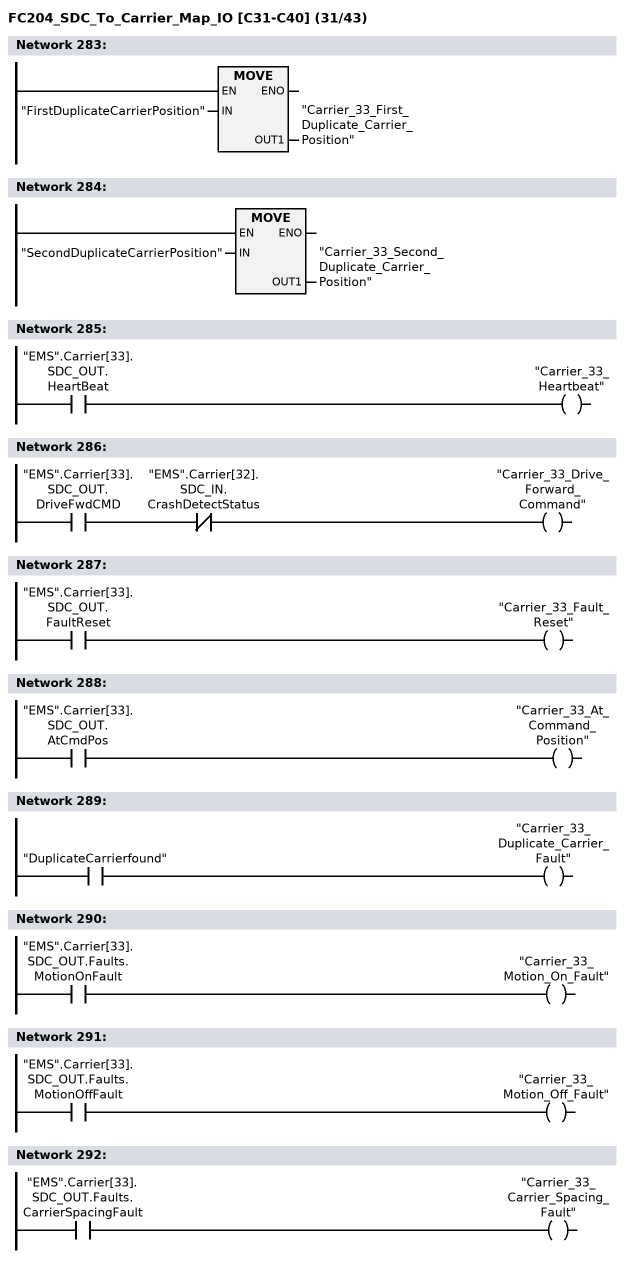
   RUNG wire#powerrail
      Move(in := "FirstDuplicateCarrierPosition", out1 => "Carrier_33_First_Duplicate_Carrier_Position")
   END_RUNG
   // the same network as SCL:
   "Carrier_33_First_Duplicate_Carrier_Position" := "FirstDuplicateCarrierPosition";
END_REGION

REGION Network 284
   RUNG wire#powerrail
      Move(in := "SecondDuplicateCarrierPosition", out1 => "Carrier_33_Second_Duplicate_Carrier_Position")
   END_RUNG
   // the same network as SCL:
   "Carrier_33_Second_Duplicate_Carrier_Position" := "SecondDuplicateCarrierPosition";
END_REGION

REGION Network 285
   RUNG wire#powerrail
      Contact( "EMS".Carrier[33].SDC_OUT.HeartBeat )
      Coil( "Carrier_33_Heartbeat" )
   END_RUNG
   // the same network as SCL:
   "Carrier_33_Heartbeat" := "EMS".Carrier[33].SDC_OUT.HeartBeat;
END_REGION

REGION Network 286
   RUNG wire#powerrail
      Contact( "EMS".Carrier[33].SDC_OUT.DriveFwdCMD )
      I_Contact( "EMS".Carrier[32].SDC_IN.CrashDetectStatus )
      Coil( "Carrier_33_Drive_Forward_Command" )
   END_RUNG
   // the same network as SCL:
   "Carrier_33_Drive_Forward_Command" := "EMS".Carrier[33].SDC_OUT.DriveFwdCMD AND NOT "EMS".Carrier[32].SDC_IN.CrashDetectStatus;
END_REGION

REGION Network 287
   RUNG wire#powerrail
      Contact( "EMS".Carrier[33].SDC_OUT.FaultReset )
      Coil( "Carrier_33_Fault_Reset" )
   END_RUNG
   // the same network as SCL:
   "Carrier_33_Fault_Reset" := "EMS".Carrier[33].SDC_OUT.FaultReset;
END_REGION

REGION Network 288
   RUNG wire#powerrail
      Contact( "EMS".Carrier[33].SDC_OUT.AtCmdPos )
      Coil( "Carrier_33_At_Command_Position" )
   END_RUNG
   // the same network as SCL:
   "Carrier_33_At_Command_Position" := "EMS".Carrier[33].SDC_OUT.AtCmdPos;
END_REGION

REGION Network 289
   RUNG wire#powerrail
      Contact( "DuplicateCarrierfound" )
      Coil( "Carrier_33_Duplicate_Carrier_Fault" )
   END_RUNG
   // the same network as SCL:
   "Carrier_33_Duplicate_Carrier_Fault" := "DuplicateCarrierfound";
END_REGION

REGION Network 290
   RUNG wire#powerrail
      Contact( "EMS".Carrier[33].SDC_OUT.Faults.MotionOnFault )
      Coil( "Carrier_33_Motion_On_Fault" )
   END_RUNG
   // the same network as SCL:
   "Carrier_33_Motion_On_Fault" := "EMS".Carrier[33].SDC_OUT.Faults.MotionOnFault;
END_REGION

REGION Network 291
   RUNG wire#powerrail
      Contact( "EMS".Carrier[33].SDC_OUT.Faults.MotionOffFault )
      Coil( "Carrier_33_Motion_Off_Fault" )
   END_RUNG
   // the same network as SCL:
   "Carrier_33_Motion_Off_Fault" := "EMS".Carrier[33].SDC_OUT.Faults.MotionOffFault;
END_REGION

REGION Network 292
   RUNG wire#powerrail
      Contact( "EMS".Carrier[33].SDC_OUT.Faults.CarrierSpacingFault )
      Coil( "Carrier_33_Carrier_Spacing_Fault" )
   END_RUNG
   // the same network as SCL:
   "Carrier_33_Carrier_Spacing_Fault" := "EMS".Carrier[33].SDC_OUT.Faults.CarrierSpacingFault;
END_REGION

REGION Network 293
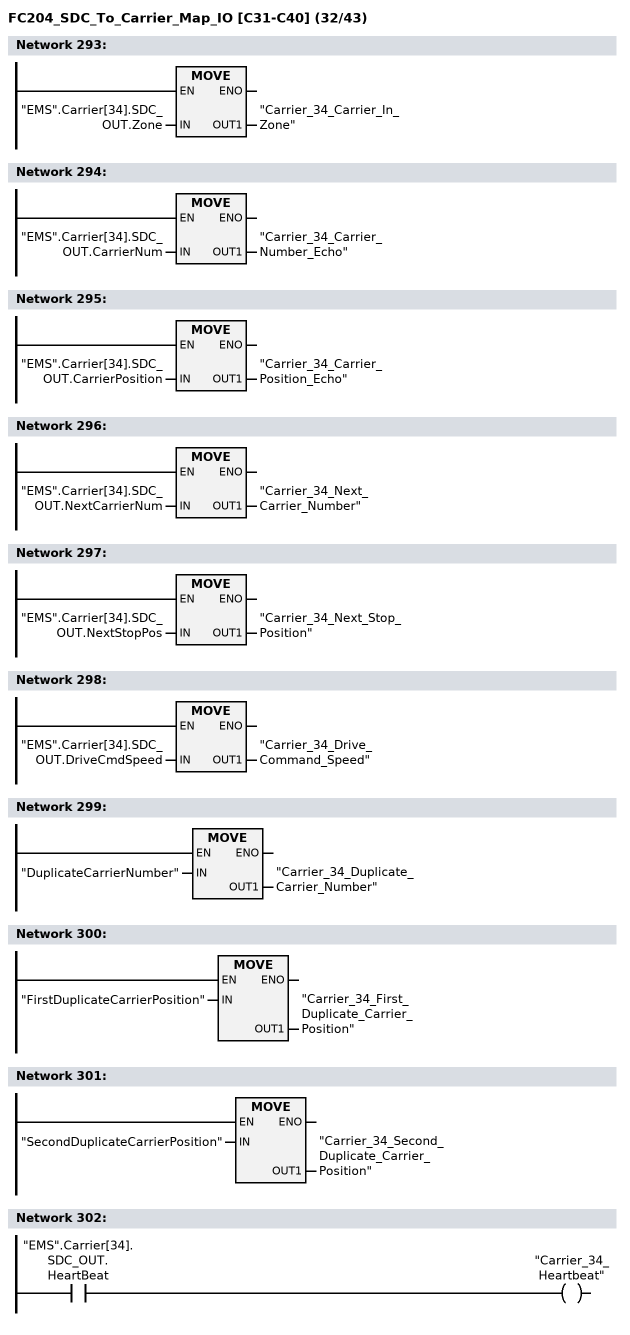
   RUNG wire#powerrail
      Move(in := "EMS".Carrier[34].SDC_OUT.Zone, out1 => "Carrier_34_Carrier_In_Zone")
   END_RUNG
   // the same network as SCL:
   "Carrier_34_Carrier_In_Zone" := "EMS".Carrier[34].SDC_OUT.Zone;
END_REGION

REGION Network 294
   RUNG wire#powerrail
      Move(in := "EMS".Carrier[34].SDC_OUT.CarrierNum, out1 => "Carrier_34_Carrier_Number_Echo")
   END_RUNG
   // the same network as SCL:
   "Carrier_34_Carrier_Number_Echo" := "EMS".Carrier[34].SDC_OUT.CarrierNum;
END_REGION

REGION Network 295
   RUNG wire#powerrail
      Move(in := "EMS".Carrier[34].SDC_OUT.CarrierPosition, out1 => "Carrier_34_Carrier_Position_Echo")
   END_RUNG
   // the same network as SCL:
   "Carrier_34_Carrier_Position_Echo" := "EMS".Carrier[34].SDC_OUT.CarrierPosition;
END_REGION

REGION Network 296
   RUNG wire#powerrail
      Move(in := "EMS".Carrier[34].SDC_OUT.NextCarrierNum, out1 => "Carrier_34_Next_Carrier_Number")
   END_RUNG
   // the same network as SCL:
   "Carrier_34_Next_Carrier_Number" := "EMS".Carrier[34].SDC_OUT.NextCarrierNum;
END_REGION

REGION Network 297
   RUNG wire#powerrail
      Move(in := "EMS".Carrier[34].SDC_OUT.NextStopPos, out1 => "Carrier_34_Next_Stop_Position")
   END_RUNG
   // the same network as SCL:
   "Carrier_34_Next_Stop_Position" := "EMS".Carrier[34].SDC_OUT.NextStopPos;
END_REGION

REGION Network 298
   RUNG wire#powerrail
      Move(in := "EMS".Carrier[34].SDC_OUT.DriveCmdSpeed, out1 => "Carrier_34_Drive_Command_Speed")
   END_RUNG
   // the same network as SCL:
   "Carrier_34_Drive_Command_Speed" := "EMS".Carrier[34].SDC_OUT.DriveCmdSpeed;
END_REGION

REGION Network 299
   RUNG wire#powerrail
      Move(in := "DuplicateCarrierNumber", out1 => "Carrier_34_Duplicate_Carrier_Number")
   END_RUNG
   // the same network as SCL:
   "Carrier_34_Duplicate_Carrier_Number" := "DuplicateCarrierNumber";
END_REGION

REGION Network 300
   RUNG wire#powerrail
      Move(in := "FirstDuplicateCarrierPosition", out1 => "Carrier_34_First_Duplicate_Carrier_Position")
   END_RUNG
   // the same network as SCL:
   "Carrier_34_First_Duplicate_Carrier_Position" := "FirstDuplicateCarrierPosition";
END_REGION

REGION Network 301
   RUNG wire#powerrail
      Move(in := "SecondDuplicateCarrierPosition", out1 => "Carrier_34_Second_Duplicate_Carrier_Position")
   END_RUNG
   // the same network as SCL:
   "Carrier_34_Second_Duplicate_Carrier_Position" := "SecondDuplicateCarrierPosition";
END_REGION

REGION Network 302
   RUNG wire#powerrail
      Contact( "EMS".Carrier[34].SDC_OUT.HeartBeat )
      Coil( "Carrier_34_Heartbeat" )
   END_RUNG
   // the same network as SCL:
   "Carrier_34_Heartbeat" := "EMS".Carrier[34].SDC_OUT.HeartBeat;
END_REGION

REGION Network 303
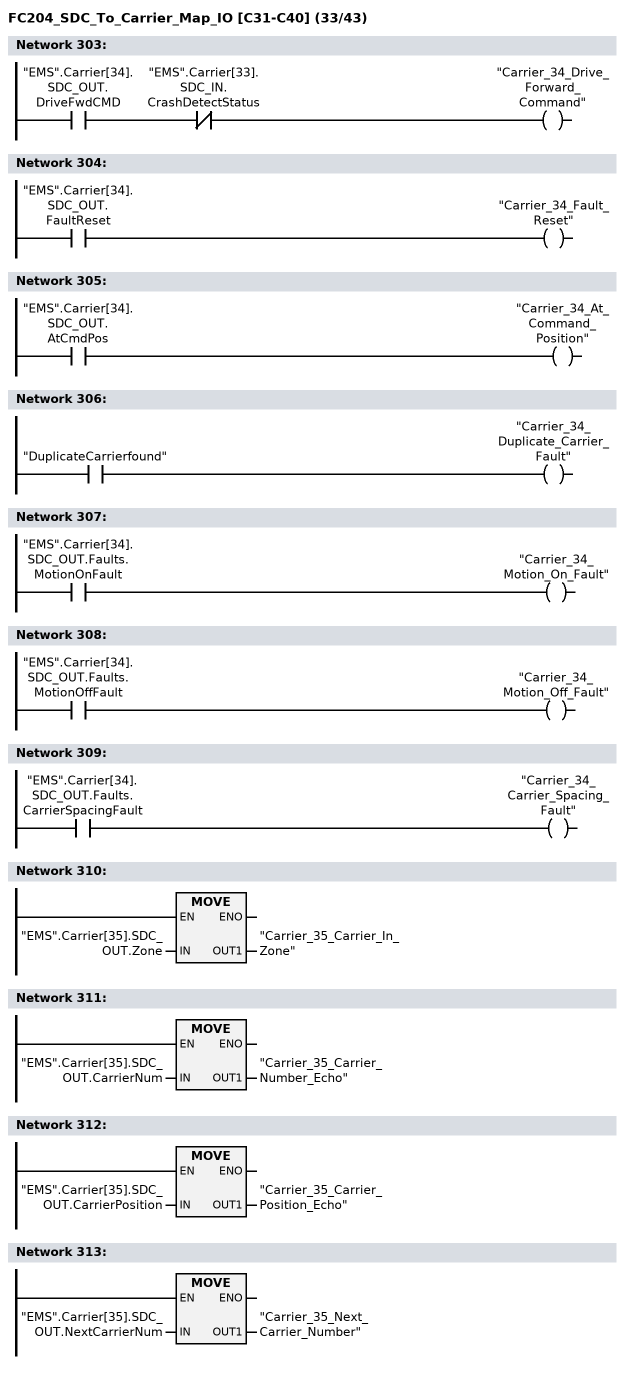
   RUNG wire#powerrail
      Contact( "EMS".Carrier[34].SDC_OUT.DriveFwdCMD )
      I_Contact( "EMS".Carrier[33].SDC_IN.CrashDetectStatus )
      Coil( "Carrier_34_Drive_Forward_Command" )
   END_RUNG
   // the same network as SCL:
   "Carrier_34_Drive_Forward_Command" := "EMS".Carrier[34].SDC_OUT.DriveFwdCMD AND NOT "EMS".Carrier[33].SDC_IN.CrashDetectStatus;
END_REGION

REGION Network 304
   RUNG wire#powerrail
      Contact( "EMS".Carrier[34].SDC_OUT.FaultReset )
      Coil( "Carrier_34_Fault_Reset" )
   END_RUNG
   // the same network as SCL:
   "Carrier_34_Fault_Reset" := "EMS".Carrier[34].SDC_OUT.FaultReset;
END_REGION

REGION Network 305
   RUNG wire#powerrail
      Contact( "EMS".Carrier[34].SDC_OUT.AtCmdPos )
      Coil( "Carrier_34_At_Command_Position" )
   END_RUNG
   // the same network as SCL:
   "Carrier_34_At_Command_Position" := "EMS".Carrier[34].SDC_OUT.AtCmdPos;
END_REGION

REGION Network 306
   RUNG wire#powerrail
      Contact( "DuplicateCarrierfound" )
      Coil( "Carrier_34_Duplicate_Carrier_Fault" )
   END_RUNG
   // the same network as SCL:
   "Carrier_34_Duplicate_Carrier_Fault" := "DuplicateCarrierfound";
END_REGION

REGION Network 307
   RUNG wire#powerrail
      Contact( "EMS".Carrier[34].SDC_OUT.Faults.MotionOnFault )
      Coil( "Carrier_34_Motion_On_Fault" )
   END_RUNG
   // the same network as SCL:
   "Carrier_34_Motion_On_Fault" := "EMS".Carrier[34].SDC_OUT.Faults.MotionOnFault;
END_REGION

REGION Network 308
   RUNG wire#powerrail
      Contact( "EMS".Carrier[34].SDC_OUT.Faults.MotionOffFault )
      Coil( "Carrier_34_Motion_Off_Fault" )
   END_RUNG
   // the same network as SCL:
   "Carrier_34_Motion_Off_Fault" := "EMS".Carrier[34].SDC_OUT.Faults.MotionOffFault;
END_REGION

REGION Network 309
   RUNG wire#powerrail
      Contact( "EMS".Carrier[34].SDC_OUT.Faults.CarrierSpacingFault )
      Coil( "Carrier_34_Carrier_Spacing_Fault" )
   END_RUNG
   // the same network as SCL:
   "Carrier_34_Carrier_Spacing_Fault" := "EMS".Carrier[34].SDC_OUT.Faults.CarrierSpacingFault;
END_REGION

REGION Network 310
   RUNG wire#powerrail
      Move(in := "EMS".Carrier[35].SDC_OUT.Zone, out1 => "Carrier_35_Carrier_In_Zone")
   END_RUNG
   // the same network as SCL:
   "Carrier_35_Carrier_In_Zone" := "EMS".Carrier[35].SDC_OUT.Zone;
END_REGION

REGION Network 311
   RUNG wire#powerrail
      Move(in := "EMS".Carrier[35].SDC_OUT.CarrierNum, out1 => "Carrier_35_Carrier_Number_Echo")
   END_RUNG
   // the same network as SCL:
   "Carrier_35_Carrier_Number_Echo" := "EMS".Carrier[35].SDC_OUT.CarrierNum;
END_REGION

REGION Network 312
   RUNG wire#powerrail
      Move(in := "EMS".Carrier[35].SDC_OUT.CarrierPosition, out1 => "Carrier_35_Carrier_Position_Echo")
   END_RUNG
   // the same network as SCL:
   "Carrier_35_Carrier_Position_Echo" := "EMS".Carrier[35].SDC_OUT.CarrierPosition;
END_REGION

REGION Network 313
   RUNG wire#powerrail
      Move(in := "EMS".Carrier[35].SDC_OUT.NextCarrierNum, out1 => "Carrier_35_Next_Carrier_Number")
   END_RUNG
   // the same network as SCL:
   "Carrier_35_Next_Carrier_Number" := "EMS".Carrier[35].SDC_OUT.NextCarrierNum;
END_REGION

REGION Network 314
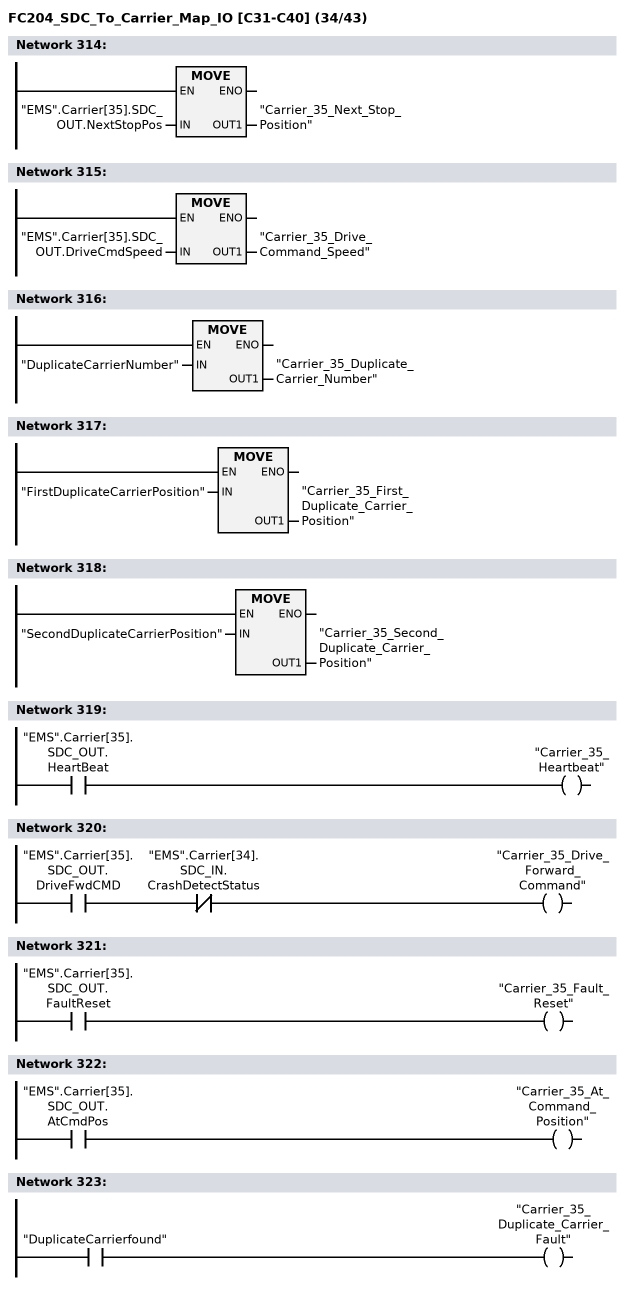
   RUNG wire#powerrail
      Move(in := "EMS".Carrier[35].SDC_OUT.NextStopPos, out1 => "Carrier_35_Next_Stop_Position")
   END_RUNG
   // the same network as SCL:
   "Carrier_35_Next_Stop_Position" := "EMS".Carrier[35].SDC_OUT.NextStopPos;
END_REGION

REGION Network 315
   RUNG wire#powerrail
      Move(in := "EMS".Carrier[35].SDC_OUT.DriveCmdSpeed, out1 => "Carrier_35_Drive_Command_Speed")
   END_RUNG
   // the same network as SCL:
   "Carrier_35_Drive_Command_Speed" := "EMS".Carrier[35].SDC_OUT.DriveCmdSpeed;
END_REGION

REGION Network 316
   RUNG wire#powerrail
      Move(in := "DuplicateCarrierNumber", out1 => "Carrier_35_Duplicate_Carrier_Number")
   END_RUNG
   // the same network as SCL:
   "Carrier_35_Duplicate_Carrier_Number" := "DuplicateCarrierNumber";
END_REGION

REGION Network 317
   RUNG wire#powerrail
      Move(in := "FirstDuplicateCarrierPosition", out1 => "Carrier_35_First_Duplicate_Carrier_Position")
   END_RUNG
   // the same network as SCL:
   "Carrier_35_First_Duplicate_Carrier_Position" := "FirstDuplicateCarrierPosition";
END_REGION

REGION Network 318
   RUNG wire#powerrail
      Move(in := "SecondDuplicateCarrierPosition", out1 => "Carrier_35_Second_Duplicate_Carrier_Position")
   END_RUNG
   // the same network as SCL:
   "Carrier_35_Second_Duplicate_Carrier_Position" := "SecondDuplicateCarrierPosition";
END_REGION

REGION Network 319
   RUNG wire#powerrail
      Contact( "EMS".Carrier[35].SDC_OUT.HeartBeat )
      Coil( "Carrier_35_Heartbeat" )
   END_RUNG
   // the same network as SCL:
   "Carrier_35_Heartbeat" := "EMS".Carrier[35].SDC_OUT.HeartBeat;
END_REGION

REGION Network 320
   RUNG wire#powerrail
      Contact( "EMS".Carrier[35].SDC_OUT.DriveFwdCMD )
      I_Contact( "EMS".Carrier[34].SDC_IN.CrashDetectStatus )
      Coil( "Carrier_35_Drive_Forward_Command" )
   END_RUNG
   // the same network as SCL:
   "Carrier_35_Drive_Forward_Command" := "EMS".Carrier[35].SDC_OUT.DriveFwdCMD AND NOT "EMS".Carrier[34].SDC_IN.CrashDetectStatus;
END_REGION

REGION Network 321
   RUNG wire#powerrail
      Contact( "EMS".Carrier[35].SDC_OUT.FaultReset )
      Coil( "Carrier_35_Fault_Reset" )
   END_RUNG
   // the same network as SCL:
   "Carrier_35_Fault_Reset" := "EMS".Carrier[35].SDC_OUT.FaultReset;
END_REGION

REGION Network 322
   RUNG wire#powerrail
      Contact( "EMS".Carrier[35].SDC_OUT.AtCmdPos )
      Coil( "Carrier_35_At_Command_Position" )
   END_RUNG
   // the same network as SCL:
   "Carrier_35_At_Command_Position" := "EMS".Carrier[35].SDC_OUT.AtCmdPos;
END_REGION

REGION Network 323
   RUNG wire#powerrail
      Contact( "DuplicateCarrierfound" )
      Coil( "Carrier_35_Duplicate_Carrier_Fault" )
   END_RUNG
   // the same network as SCL:
   "Carrier_35_Duplicate_Carrier_Fault" := "DuplicateCarrierfound";
END_REGION

REGION Network 324
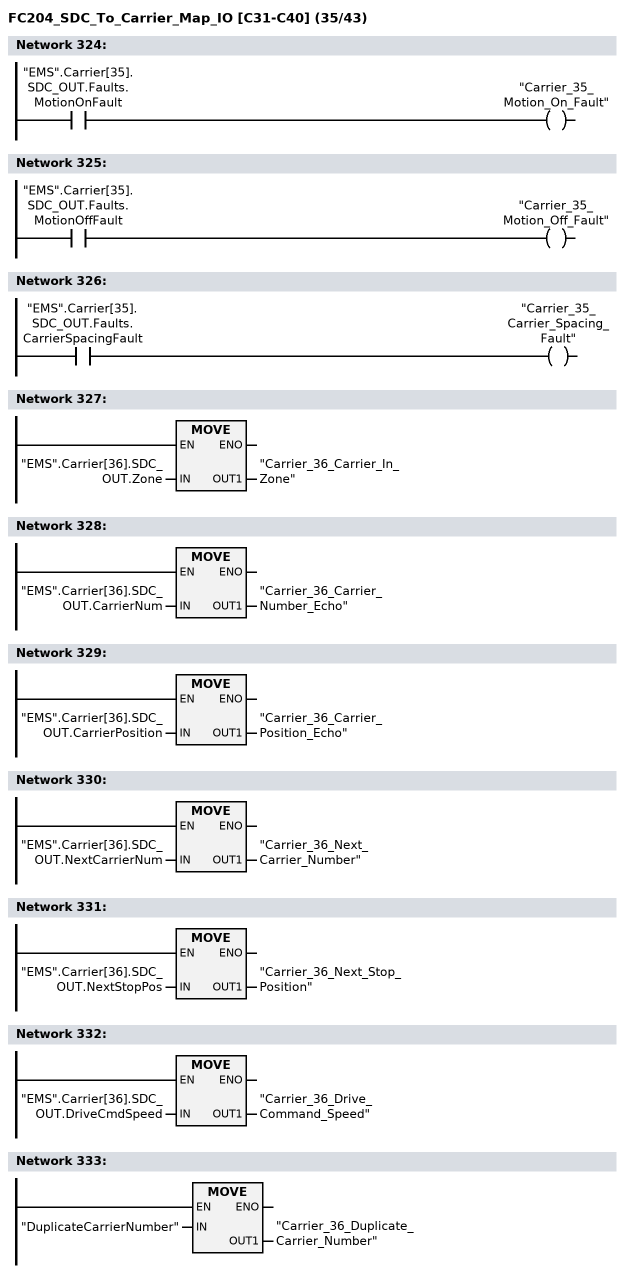
   RUNG wire#powerrail
      Contact( "EMS".Carrier[35].SDC_OUT.Faults.MotionOnFault )
      Coil( "Carrier_35_Motion_On_Fault" )
   END_RUNG
   // the same network as SCL:
   "Carrier_35_Motion_On_Fault" := "EMS".Carrier[35].SDC_OUT.Faults.MotionOnFault;
END_REGION

REGION Network 325
   RUNG wire#powerrail
      Contact( "EMS".Carrier[35].SDC_OUT.Faults.MotionOffFault )
      Coil( "Carrier_35_Motion_Off_Fault" )
   END_RUNG
   // the same network as SCL:
   "Carrier_35_Motion_Off_Fault" := "EMS".Carrier[35].SDC_OUT.Faults.MotionOffFault;
END_REGION

REGION Network 326
   RUNG wire#powerrail
      Contact( "EMS".Carrier[35].SDC_OUT.Faults.CarrierSpacingFault )
      Coil( "Carrier_35_Carrier_Spacing_Fault" )
   END_RUNG
   // the same network as SCL:
   "Carrier_35_Carrier_Spacing_Fault" := "EMS".Carrier[35].SDC_OUT.Faults.CarrierSpacingFault;
END_REGION

REGION Network 327
   RUNG wire#powerrail
      Move(in := "EMS".Carrier[36].SDC_OUT.Zone, out1 => "Carrier_36_Carrier_In_Zone")
   END_RUNG
   // the same network as SCL:
   "Carrier_36_Carrier_In_Zone" := "EMS".Carrier[36].SDC_OUT.Zone;
END_REGION

REGION Network 328
   RUNG wire#powerrail
      Move(in := "EMS".Carrier[36].SDC_OUT.CarrierNum, out1 => "Carrier_36_Carrier_Number_Echo")
   END_RUNG
   // the same network as SCL:
   "Carrier_36_Carrier_Number_Echo" := "EMS".Carrier[36].SDC_OUT.CarrierNum;
END_REGION

REGION Network 329
   RUNG wire#powerrail
      Move(in := "EMS".Carrier[36].SDC_OUT.CarrierPosition, out1 => "Carrier_36_Carrier_Position_Echo")
   END_RUNG
   // the same network as SCL:
   "Carrier_36_Carrier_Position_Echo" := "EMS".Carrier[36].SDC_OUT.CarrierPosition;
END_REGION

REGION Network 330
   RUNG wire#powerrail
      Move(in := "EMS".Carrier[36].SDC_OUT.NextCarrierNum, out1 => "Carrier_36_Next_Carrier_Number")
   END_RUNG
   // the same network as SCL:
   "Carrier_36_Next_Carrier_Number" := "EMS".Carrier[36].SDC_OUT.NextCarrierNum;
END_REGION

REGION Network 331
   RUNG wire#powerrail
      Move(in := "EMS".Carrier[36].SDC_OUT.NextStopPos, out1 => "Carrier_36_Next_Stop_Position")
   END_RUNG
   // the same network as SCL:
   "Carrier_36_Next_Stop_Position" := "EMS".Carrier[36].SDC_OUT.NextStopPos;
END_REGION

REGION Network 332
   RUNG wire#powerrail
      Move(in := "EMS".Carrier[36].SDC_OUT.DriveCmdSpeed, out1 => "Carrier_36_Drive_Command_Speed")
   END_RUNG
   // the same network as SCL:
   "Carrier_36_Drive_Command_Speed" := "EMS".Carrier[36].SDC_OUT.DriveCmdSpeed;
END_REGION

REGION Network 333
   RUNG wire#powerrail
      Move(in := "DuplicateCarrierNumber", out1 => "Carrier_36_Duplicate_Carrier_Number")
   END_RUNG
   // the same network as SCL:
   "Carrier_36_Duplicate_Carrier_Number" := "DuplicateCarrierNumber";
END_REGION

REGION Network 334
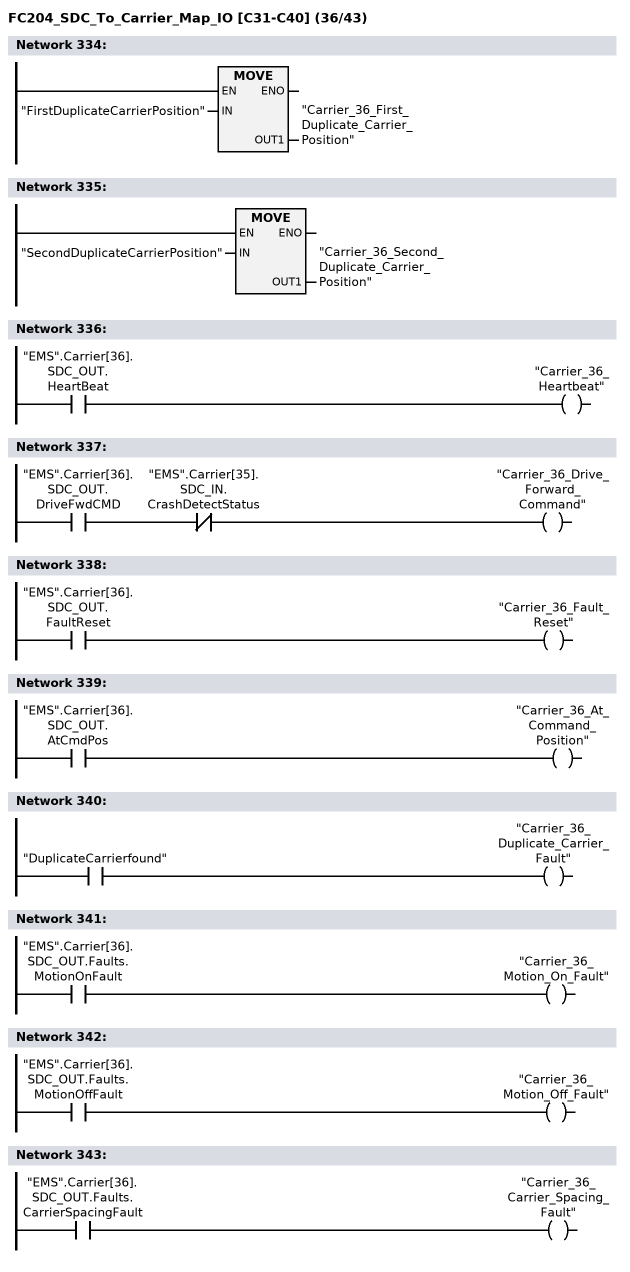
   RUNG wire#powerrail
      Move(in := "FirstDuplicateCarrierPosition", out1 => "Carrier_36_First_Duplicate_Carrier_Position")
   END_RUNG
   // the same network as SCL:
   "Carrier_36_First_Duplicate_Carrier_Position" := "FirstDuplicateCarrierPosition";
END_REGION

REGION Network 335
   RUNG wire#powerrail
      Move(in := "SecondDuplicateCarrierPosition", out1 => "Carrier_36_Second_Duplicate_Carrier_Position")
   END_RUNG
   // the same network as SCL:
   "Carrier_36_Second_Duplicate_Carrier_Position" := "SecondDuplicateCarrierPosition";
END_REGION

REGION Network 336
   RUNG wire#powerrail
      Contact( "EMS".Carrier[36].SDC_OUT.HeartBeat )
      Coil( "Carrier_36_Heartbeat" )
   END_RUNG
   // the same network as SCL:
   "Carrier_36_Heartbeat" := "EMS".Carrier[36].SDC_OUT.HeartBeat;
END_REGION

REGION Network 337
   RUNG wire#powerrail
      Contact( "EMS".Carrier[36].SDC_OUT.DriveFwdCMD )
      I_Contact( "EMS".Carrier[35].SDC_IN.CrashDetectStatus )
      Coil( "Carrier_36_Drive_Forward_Command" )
   END_RUNG
   // the same network as SCL:
   "Carrier_36_Drive_Forward_Command" := "EMS".Carrier[36].SDC_OUT.DriveFwdCMD AND NOT "EMS".Carrier[35].SDC_IN.CrashDetectStatus;
END_REGION

REGION Network 338
   RUNG wire#powerrail
      Contact( "EMS".Carrier[36].SDC_OUT.FaultReset )
      Coil( "Carrier_36_Fault_Reset" )
   END_RUNG
   // the same network as SCL:
   "Carrier_36_Fault_Reset" := "EMS".Carrier[36].SDC_OUT.FaultReset;
END_REGION

REGION Network 339
   RUNG wire#powerrail
      Contact( "EMS".Carrier[36].SDC_OUT.AtCmdPos )
      Coil( "Carrier_36_At_Command_Position" )
   END_RUNG
   // the same network as SCL:
   "Carrier_36_At_Command_Position" := "EMS".Carrier[36].SDC_OUT.AtCmdPos;
END_REGION

REGION Network 340
   RUNG wire#powerrail
      Contact( "DuplicateCarrierfound" )
      Coil( "Carrier_36_Duplicate_Carrier_Fault" )
   END_RUNG
   // the same network as SCL:
   "Carrier_36_Duplicate_Carrier_Fault" := "DuplicateCarrierfound";
END_REGION

REGION Network 341
   RUNG wire#powerrail
      Contact( "EMS".Carrier[36].SDC_OUT.Faults.MotionOnFault )
      Coil( "Carrier_36_Motion_On_Fault" )
   END_RUNG
   // the same network as SCL:
   "Carrier_36_Motion_On_Fault" := "EMS".Carrier[36].SDC_OUT.Faults.MotionOnFault;
END_REGION

REGION Network 342
   RUNG wire#powerrail
      Contact( "EMS".Carrier[36].SDC_OUT.Faults.MotionOffFault )
      Coil( "Carrier_36_Motion_Off_Fault" )
   END_RUNG
   // the same network as SCL:
   "Carrier_36_Motion_Off_Fault" := "EMS".Carrier[36].SDC_OUT.Faults.MotionOffFault;
END_REGION

REGION Network 343
   RUNG wire#powerrail
      Contact( "EMS".Carrier[36].SDC_OUT.Faults.CarrierSpacingFault )
      Coil( "Carrier_36_Carrier_Spacing_Fault" )
   END_RUNG
   // the same network as SCL:
   "Carrier_36_Carrier_Spacing_Fault" := "EMS".Carrier[36].SDC_OUT.Faults.CarrierSpacingFault;
END_REGION

REGION Network 344
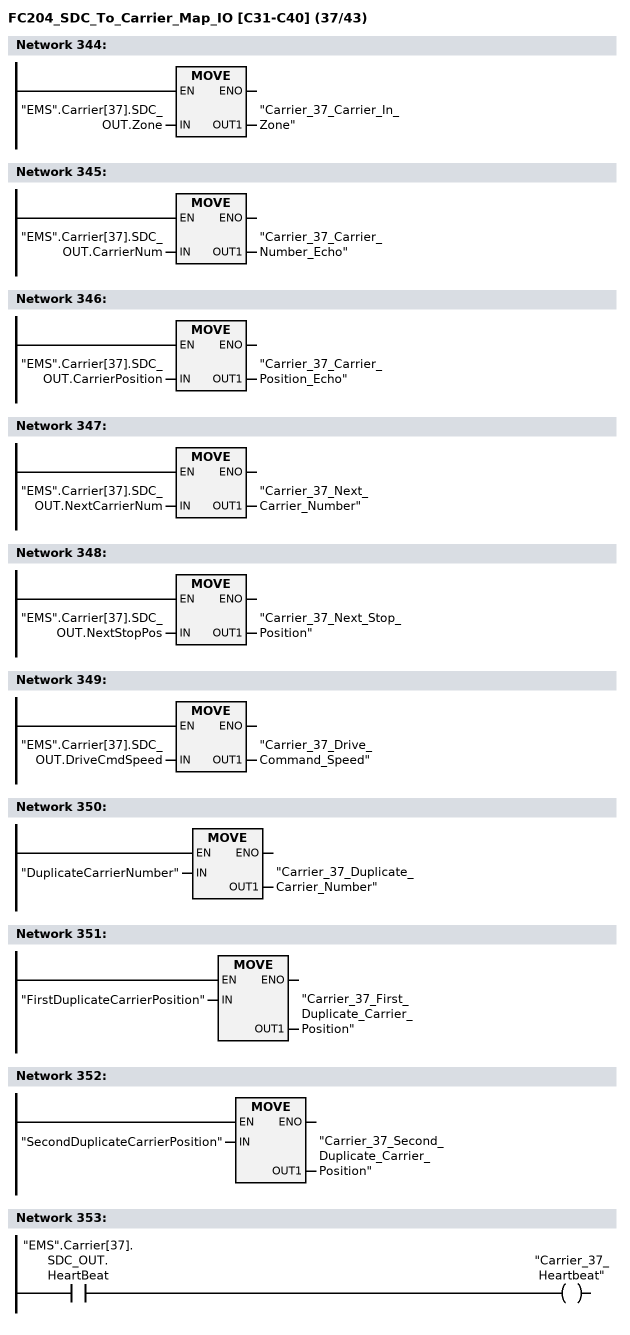
   RUNG wire#powerrail
      Move(in := "EMS".Carrier[37].SDC_OUT.Zone, out1 => "Carrier_37_Carrier_In_Zone")
   END_RUNG
   // the same network as SCL:
   "Carrier_37_Carrier_In_Zone" := "EMS".Carrier[37].SDC_OUT.Zone;
END_REGION

REGION Network 345
   RUNG wire#powerrail
      Move(in := "EMS".Carrier[37].SDC_OUT.CarrierNum, out1 => "Carrier_37_Carrier_Number_Echo")
   END_RUNG
   // the same network as SCL:
   "Carrier_37_Carrier_Number_Echo" := "EMS".Carrier[37].SDC_OUT.CarrierNum;
END_REGION

REGION Network 346
   RUNG wire#powerrail
      Move(in := "EMS".Carrier[37].SDC_OUT.CarrierPosition, out1 => "Carrier_37_Carrier_Position_Echo")
   END_RUNG
   // the same network as SCL:
   "Carrier_37_Carrier_Position_Echo" := "EMS".Carrier[37].SDC_OUT.CarrierPosition;
END_REGION

REGION Network 347
   RUNG wire#powerrail
      Move(in := "EMS".Carrier[37].SDC_OUT.NextCarrierNum, out1 => "Carrier_37_Next_Carrier_Number")
   END_RUNG
   // the same network as SCL:
   "Carrier_37_Next_Carrier_Number" := "EMS".Carrier[37].SDC_OUT.NextCarrierNum;
END_REGION

REGION Network 348
   RUNG wire#powerrail
      Move(in := "EMS".Carrier[37].SDC_OUT.NextStopPos, out1 => "Carrier_37_Next_Stop_Position")
   END_RUNG
   // the same network as SCL:
   "Carrier_37_Next_Stop_Position" := "EMS".Carrier[37].SDC_OUT.NextStopPos;
END_REGION

REGION Network 349
   RUNG wire#powerrail
      Move(in := "EMS".Carrier[37].SDC_OUT.DriveCmdSpeed, out1 => "Carrier_37_Drive_Command_Speed")
   END_RUNG
   // the same network as SCL:
   "Carrier_37_Drive_Command_Speed" := "EMS".Carrier[37].SDC_OUT.DriveCmdSpeed;
END_REGION

REGION Network 350
   RUNG wire#powerrail
      Move(in := "DuplicateCarrierNumber", out1 => "Carrier_37_Duplicate_Carrier_Number")
   END_RUNG
   // the same network as SCL:
   "Carrier_37_Duplicate_Carrier_Number" := "DuplicateCarrierNumber";
END_REGION

REGION Network 351
   RUNG wire#powerrail
      Move(in := "FirstDuplicateCarrierPosition", out1 => "Carrier_37_First_Duplicate_Carrier_Position")
   END_RUNG
   // the same network as SCL:
   "Carrier_37_First_Duplicate_Carrier_Position" := "FirstDuplicateCarrierPosition";
END_REGION

REGION Network 352
   RUNG wire#powerrail
      Move(in := "SecondDuplicateCarrierPosition", out1 => "Carrier_37_Second_Duplicate_Carrier_Position")
   END_RUNG
   // the same network as SCL:
   "Carrier_37_Second_Duplicate_Carrier_Position" := "SecondDuplicateCarrierPosition";
END_REGION

REGION Network 353
   RUNG wire#powerrail
      Contact( "EMS".Carrier[37].SDC_OUT.HeartBeat )
      Coil( "Carrier_37_Heartbeat" )
   END_RUNG
   // the same network as SCL:
   "Carrier_37_Heartbeat" := "EMS".Carrier[37].SDC_OUT.HeartBeat;
END_REGION

REGION Network 354
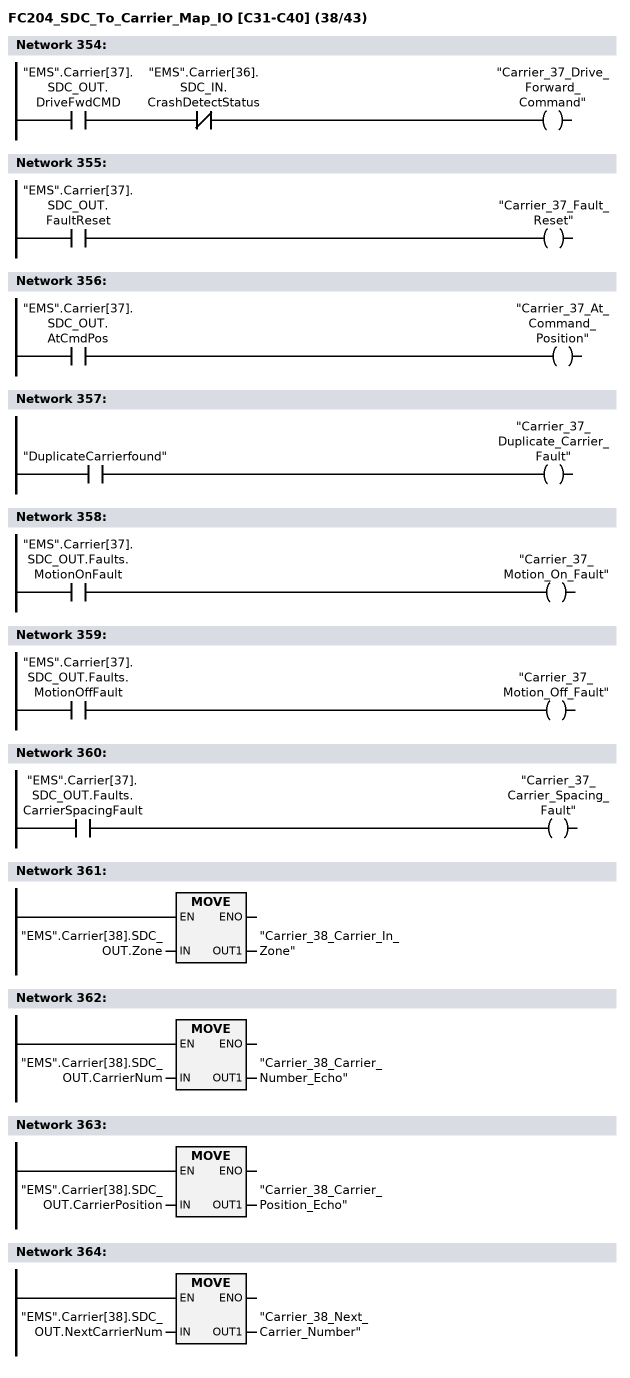
   RUNG wire#powerrail
      Contact( "EMS".Carrier[37].SDC_OUT.DriveFwdCMD )
      I_Contact( "EMS".Carrier[36].SDC_IN.CrashDetectStatus )
      Coil( "Carrier_37_Drive_Forward_Command" )
   END_RUNG
   // the same network as SCL:
   "Carrier_37_Drive_Forward_Command" := "EMS".Carrier[37].SDC_OUT.DriveFwdCMD AND NOT "EMS".Carrier[36].SDC_IN.CrashDetectStatus;
END_REGION

REGION Network 355
   RUNG wire#powerrail
      Contact( "EMS".Carrier[37].SDC_OUT.FaultReset )
      Coil( "Carrier_37_Fault_Reset" )
   END_RUNG
   // the same network as SCL:
   "Carrier_37_Fault_Reset" := "EMS".Carrier[37].SDC_OUT.FaultReset;
END_REGION

REGION Network 356
   RUNG wire#powerrail
      Contact( "EMS".Carrier[37].SDC_OUT.AtCmdPos )
      Coil( "Carrier_37_At_Command_Position" )
   END_RUNG
   // the same network as SCL:
   "Carrier_37_At_Command_Position" := "EMS".Carrier[37].SDC_OUT.AtCmdPos;
END_REGION

REGION Network 357
   RUNG wire#powerrail
      Contact( "DuplicateCarrierfound" )
      Coil( "Carrier_37_Duplicate_Carrier_Fault" )
   END_RUNG
   // the same network as SCL:
   "Carrier_37_Duplicate_Carrier_Fault" := "DuplicateCarrierfound";
END_REGION

REGION Network 358
   RUNG wire#powerrail
      Contact( "EMS".Carrier[37].SDC_OUT.Faults.MotionOnFault )
      Coil( "Carrier_37_Motion_On_Fault" )
   END_RUNG
   // the same network as SCL:
   "Carrier_37_Motion_On_Fault" := "EMS".Carrier[37].SDC_OUT.Faults.MotionOnFault;
END_REGION

REGION Network 359
   RUNG wire#powerrail
      Contact( "EMS".Carrier[37].SDC_OUT.Faults.MotionOffFault )
      Coil( "Carrier_37_Motion_Off_Fault" )
   END_RUNG
   // the same network as SCL:
   "Carrier_37_Motion_Off_Fault" := "EMS".Carrier[37].SDC_OUT.Faults.MotionOffFault;
END_REGION

REGION Network 360
   RUNG wire#powerrail
      Contact( "EMS".Carrier[37].SDC_OUT.Faults.CarrierSpacingFault )
      Coil( "Carrier_37_Carrier_Spacing_Fault" )
   END_RUNG
   // the same network as SCL:
   "Carrier_37_Carrier_Spacing_Fault" := "EMS".Carrier[37].SDC_OUT.Faults.CarrierSpacingFault;
END_REGION

REGION Network 361
   RUNG wire#powerrail
      Move(in := "EMS".Carrier[38].SDC_OUT.Zone, out1 => "Carrier_38_Carrier_In_Zone")
   END_RUNG
   // the same network as SCL:
   "Carrier_38_Carrier_In_Zone" := "EMS".Carrier[38].SDC_OUT.Zone;
END_REGION

REGION Network 362
   RUNG wire#powerrail
      Move(in := "EMS".Carrier[38].SDC_OUT.CarrierNum, out1 => "Carrier_38_Carrier_Number_Echo")
   END_RUNG
   // the same network as SCL:
   "Carrier_38_Carrier_Number_Echo" := "EMS".Carrier[38].SDC_OUT.CarrierNum;
END_REGION

REGION Network 363
   RUNG wire#powerrail
      Move(in := "EMS".Carrier[38].SDC_OUT.CarrierPosition, out1 => "Carrier_38_Carrier_Position_Echo")
   END_RUNG
   // the same network as SCL:
   "Carrier_38_Carrier_Position_Echo" := "EMS".Carrier[38].SDC_OUT.CarrierPosition;
END_REGION

REGION Network 364
   RUNG wire#powerrail
      Move(in := "EMS".Carrier[38].SDC_OUT.NextCarrierNum, out1 => "Carrier_38_Next_Carrier_Number")
   END_RUNG
   // the same network as SCL:
   "Carrier_38_Next_Carrier_Number" := "EMS".Carrier[38].SDC_OUT.NextCarrierNum;
END_REGION

REGION Network 365
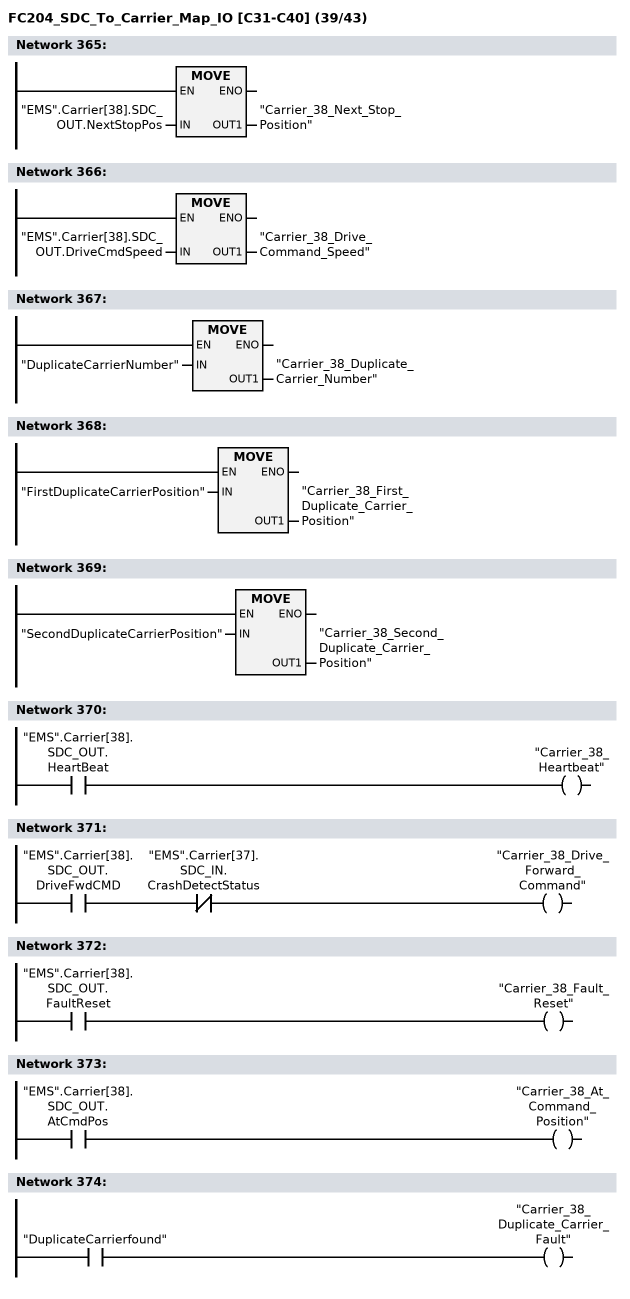
   RUNG wire#powerrail
      Move(in := "EMS".Carrier[38].SDC_OUT.NextStopPos, out1 => "Carrier_38_Next_Stop_Position")
   END_RUNG
   // the same network as SCL:
   "Carrier_38_Next_Stop_Position" := "EMS".Carrier[38].SDC_OUT.NextStopPos;
END_REGION

REGION Network 366
   RUNG wire#powerrail
      Move(in := "EMS".Carrier[38].SDC_OUT.DriveCmdSpeed, out1 => "Carrier_38_Drive_Command_Speed")
   END_RUNG
   // the same network as SCL:
   "Carrier_38_Drive_Command_Speed" := "EMS".Carrier[38].SDC_OUT.DriveCmdSpeed;
END_REGION

REGION Network 367
   RUNG wire#powerrail
      Move(in := "DuplicateCarrierNumber", out1 => "Carrier_38_Duplicate_Carrier_Number")
   END_RUNG
   // the same network as SCL:
   "Carrier_38_Duplicate_Carrier_Number" := "DuplicateCarrierNumber";
END_REGION

REGION Network 368
   RUNG wire#powerrail
      Move(in := "FirstDuplicateCarrierPosition", out1 => "Carrier_38_First_Duplicate_Carrier_Position")
   END_RUNG
   // the same network as SCL:
   "Carrier_38_First_Duplicate_Carrier_Position" := "FirstDuplicateCarrierPosition";
END_REGION

REGION Network 369
   RUNG wire#powerrail
      Move(in := "SecondDuplicateCarrierPosition", out1 => "Carrier_38_Second_Duplicate_Carrier_Position")
   END_RUNG
   // the same network as SCL:
   "Carrier_38_Second_Duplicate_Carrier_Position" := "SecondDuplicateCarrierPosition";
END_REGION

REGION Network 370
   RUNG wire#powerrail
      Contact( "EMS".Carrier[38].SDC_OUT.HeartBeat )
      Coil( "Carrier_38_Heartbeat" )
   END_RUNG
   // the same network as SCL:
   "Carrier_38_Heartbeat" := "EMS".Carrier[38].SDC_OUT.HeartBeat;
END_REGION

REGION Network 371
   RUNG wire#powerrail
      Contact( "EMS".Carrier[38].SDC_OUT.DriveFwdCMD )
      I_Contact( "EMS".Carrier[37].SDC_IN.CrashDetectStatus )
      Coil( "Carrier_38_Drive_Forward_Command" )
   END_RUNG
   // the same network as SCL:
   "Carrier_38_Drive_Forward_Command" := "EMS".Carrier[38].SDC_OUT.DriveFwdCMD AND NOT "EMS".Carrier[37].SDC_IN.CrashDetectStatus;
END_REGION

REGION Network 372
   RUNG wire#powerrail
      Contact( "EMS".Carrier[38].SDC_OUT.FaultReset )
      Coil( "Carrier_38_Fault_Reset" )
   END_RUNG
   // the same network as SCL:
   "Carrier_38_Fault_Reset" := "EMS".Carrier[38].SDC_OUT.FaultReset;
END_REGION

REGION Network 373
   RUNG wire#powerrail
      Contact( "EMS".Carrier[38].SDC_OUT.AtCmdPos )
      Coil( "Carrier_38_At_Command_Position" )
   END_RUNG
   // the same network as SCL:
   "Carrier_38_At_Command_Position" := "EMS".Carrier[38].SDC_OUT.AtCmdPos;
END_REGION

REGION Network 374
   RUNG wire#powerrail
      Contact( "DuplicateCarrierfound" )
      Coil( "Carrier_38_Duplicate_Carrier_Fault" )
   END_RUNG
   // the same network as SCL:
   "Carrier_38_Duplicate_Carrier_Fault" := "DuplicateCarrierfound";
END_REGION

REGION Network 375
